// TIA Portal project "MCP_RB001002" (V15.1) (continued)
   SendWChar[1891] := WCHAR#' ';
   SendWChar[1892] := WCHAR#' ';
   SendWChar[1893] := WCHAR#' ';
   SendWChar[1894] := WCHAR#' ';
   SendWChar[1895] := WCHAR#' ';
   SendWChar[1896] := WCHAR#' ';
   SendWChar[1897] := WCHAR#' ';
   SendWChar[1898] := WCHAR#' ';
   SendWChar[1899] := WCHAR#' ';
   SendWChar[1900] := WCHAR#' ';
   SendWChar[1901] := WCHAR#' ';
   SendWChar[1902] := WCHAR#' ';
   SendWChar[1903] := WCHAR#' ';
   SendWChar[1904] := WCHAR#' ';
   SendWChar[1905] := WCHAR#' ';
   SendWChar[1906] := WCHAR#' ';
   SendWChar[1907] := WCHAR#' ';
   SendWChar[1908] := WCHAR#' ';
   SendWChar[1909] := WCHAR#' ';
   SendWChar[1910] := WCHAR#' ';
   SendWChar[1911] := WCHAR#' ';
   SendWChar[1912] := WCHAR#' ';
   SendWChar[1913] := WCHAR#' ';
   SendWChar[1914] := WCHAR#' ';
   SendWChar[1915] := WCHAR#' ';
   SendWChar[1916] := WCHAR#' ';
   SendWChar[1917] := WCHAR#' ';
   SendWChar[1918] := WCHAR#' ';
   SendWChar[1919] := WCHAR#' ';
   SendWChar[1920] := WCHAR#' ';
   SendWChar[1921] := WCHAR#' ';
   SendWChar[1922] := WCHAR#' ';
   SendWChar[1923] := WCHAR#' ';
   SendWChar[1924] := WCHAR#' ';
   SendWChar[1925] := WCHAR#' ';
   SendWChar[1926] := WCHAR#' ';
   SendWChar[1927] := WCHAR#' ';
   SendWChar[1928] := WCHAR#' ';
   SendWChar[1929] := WCHAR#' ';
   SendWChar[1930] := WCHAR#' ';
   SendWChar[1931] := WCHAR#' ';
   SendWChar[1932] := WCHAR#' ';
   SendWChar[1933] := WCHAR#' ';
   SendWChar[1934] := WCHAR#' ';
   SendWChar[1935] := WCHAR#' ';
   SendWChar[1936] := WCHAR#' ';
   SendWChar[1937] := WCHAR#' ';
   SendWChar[1938] := WCHAR#' ';
   SendWChar[1939] := WCHAR#' ';
   SendWChar[1940] := WCHAR#' ';
   SendWChar[1941] := WCHAR#' ';
   SendWChar[1942] := WCHAR#' ';
   SendWChar[1943] := WCHAR#' ';
   SendWChar[1944] := WCHAR#' ';
   SendWChar[1945] := WCHAR#' ';
   SendWChar[1946] := WCHAR#' ';
   SendWChar[1947] := WCHAR#' ';
   SendWChar[1948] := WCHAR#' ';
   SendWChar[1949] := WCHAR#' ';
   SendWChar[1950] := WCHAR#' ';
   SendWChar[1951] := WCHAR#' ';
   SendWChar[1952] := WCHAR#' ';
   SendWChar[1953] := WCHAR#' ';
   SendWChar[1954] := WCHAR#' ';
   SendWChar[1955] := WCHAR#' ';
   SendWChar[1956] := WCHAR#' ';
   SendWChar[1957] := WCHAR#' ';
   SendWChar[1958] := WCHAR#' ';
   SendWChar[1959] := WCHAR#' ';
   SendWChar[1960] := WCHAR#' ';
   SendWChar[1961] := WCHAR#' ';
   SendWChar[1962] := WCHAR#' ';
   SendWChar[1963] := WCHAR#' ';
   SendWChar[1964] := WCHAR#' ';
   SendWChar[1965] := WCHAR#' ';
   SendWChar[1966] := WCHAR#' ';
   SendWChar[1967] := WCHAR#' ';
   SendWChar[1968] := WCHAR#' ';
   SendWChar[1969] := WCHAR#' ';
   SendWChar[1970] := WCHAR#' ';
   SendWChar[1971] := WCHAR#' ';
   SendWChar[1972] := WCHAR#' ';
   SendWChar[1973] := WCHAR#' ';
   SendWChar[1974] := WCHAR#' ';
   SendWChar[1975] := WCHAR#' ';
   SendWChar[1976] := WCHAR#' ';
   SendWChar[1977] := WCHAR#' ';
   SendWChar[1978] := WCHAR#' ';
   SendWChar[1979] := WCHAR#' ';
   SendWChar[1980] := WCHAR#' ';
   SendWChar[1981] := WCHAR#' ';
   SendWChar[1982] := WCHAR#' ';
   SendWChar[1983] := WCHAR#' ';
   SendWChar[1984] := WCHAR#' ';
   SendWChar[1985] := WCHAR#' ';
   SendWChar[1986] := WCHAR#' ';
   SendWChar[1987] := WCHAR#' ';
   SendWChar[1988] := WCHAR#' ';
   SendWChar[1989] := WCHAR#' ';
   SendWChar[1990] := WCHAR#' ';
   SendWChar[1991] := WCHAR#' ';
   SendWChar[1992] := WCHAR#' ';
   SendWChar[1993] := WCHAR#' ';
   SendWChar[1994] := WCHAR#' ';
   SendWChar[1995] := WCHAR#' ';
   SendWChar[1996] := WCHAR#' ';
   SendWChar[1997] := WCHAR#' ';
   SendWChar[1998] := WCHAR#' ';
   SendWChar[1999] := WCHAR#' ';
   SendWChar[2000] := WCHAR#' ';
   SendWChar[2001] := WCHAR#' ';
   SendWChar[2002] := WCHAR#' ';
   SendWChar[2003] := WCHAR#' ';
   SendWChar[2004] := WCHAR#' ';
   SendWChar[2005] := WCHAR#' ';
   SendWChar[2006] := WCHAR#' ';
   SendWChar[2007] := WCHAR#' ';
   SendWChar[2008] := WCHAR#' ';
   SendWChar[2009] := WCHAR#' ';
   SendWChar[2010] := WCHAR#' ';
   SendWChar[2011] := WCHAR#' ';
   SendWChar[2012] := WCHAR#' ';
   SendWChar[2013] := WCHAR#' ';
   SendWChar[2014] := WCHAR#' ';
   SendWChar[2015] := WCHAR#' ';
   SendWChar[2016] := WCHAR#' ';
   SendWChar[2017] := WCHAR#' ';
   SendWChar[2018] := WCHAR#' ';
   SendWChar[2019] := WCHAR#' ';
   SendWChar[2020] := WCHAR#' ';
   SendWChar[2021] := WCHAR#' ';
   SendWChar[2022] := WCHAR#' ';
   SendWChar[2023] := WCHAR#' ';
   SendWChar[2024] := WCHAR#' ';
   SendWChar[2025] := WCHAR#' ';
   SendWChar[2026] := WCHAR#' ';
   SendWChar[2027] := WCHAR#' ';
   SendWChar[2028] := WCHAR#' ';
   SendWChar[2029] := WCHAR#' ';
   SendWChar[2030] := WCHAR#' ';
   SendWChar[2031] := WCHAR#' ';
   SendWChar[2032] := WCHAR#' ';
   SendWChar[2033] := WCHAR#' ';
   SendWChar[2034] := WCHAR#' ';
   SendWChar[2035] := WCHAR#' ';
   SendWChar[2036] := WCHAR#' ';
   SendWChar[2037] := WCHAR#' ';
   SendWChar[2038] := WCHAR#' ';
   SendWChar[2039] := WCHAR#' ';
   SendWChar[2040] := WCHAR#' ';
   SendWChar[2041] := WCHAR#' ';
   SendWChar[2042] := WCHAR#' ';
   SendWChar[2043] := WCHAR#' ';
   SendWChar[2044] := WCHAR#' ';
   SendWChar[2045] := WCHAR#' ';
   SendWChar[2046] := WCHAR#' ';
   SendWChar[2047] := WCHAR#' ';
   SendWChar[2048] := WCHAR#' ';
END_DATA_BLOCK

DATA_BLOCK "uMySQL_Use_DB"   // DB902
{ S7_Optimized_Access := 'TRUE' }
VERSION : 0.1
// stored: InstanceOfName uMySQL_Use
"uMySQL_Use"
BEGIN
END_DATA_BLOCK

DATA_BLOCK "uMySQL_Command_DB"   // DB903
{ S7_Optimized_Access := 'TRUE' }
VERSION : 0.1
// stored: InstanceOfName uMySQL_Command
"uMySQL_Command"
BEGIN
END_DATA_BLOCK

DATA_BLOCK "uMySQL_Query_DB"   // DB904
{ S7_Optimized_Access := 'TRUE' }
VERSION : 0.1
// stored: InstanceOfName uMySQL_Query
"uMySQL_Query"
BEGIN
END_DATA_BLOCK

// folder: (top level)

FUNCTION_BLOCK "温控相机解码"   // FB410, LAD
{ S7_Optimized_Access := 'TRUE' }
VERSION : 0.1
   VAR RETAIN
      Connparm : TCON_IP_v4;
   END_VAR
   VAR
      TRCV_C_Instance : TRCV_C;
      RECV_Data : Array[0..1023] of Byte;
   END_VAR
   // Connparm.InterfaceId := 64;
   // Connparm.ID := 16#65;
   // Connparm.ActiveEstablished := false;
   // Connparm.LocalPort := 9840;
BEGIN

REGION Network 1
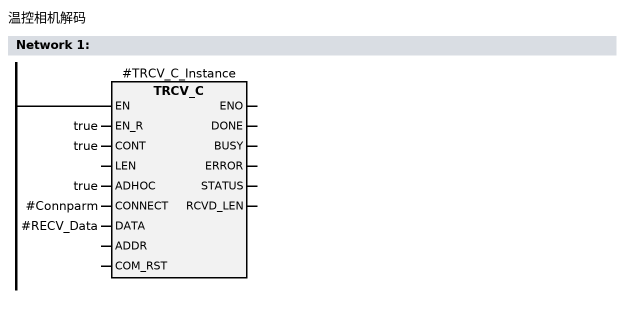
   #TRCV_C_Instance(EN_R := true, CONT := true, ADHOC := true, CONNECT := #Connparm, DATA := #RECV_Data);   // TRCV_C
END_REGION
END_FUNCTION_BLOCK

FUNCTION "精炼机数据处理" : Void   // FC100, LAD
{ S7_Optimized_Access := 'TRUE' }
VERSION : 0.1
   VAR_TEMP   // added for the SCL form of the ladder/FBD networks
      _w1 : Bool;
   END_VAR
BEGIN

REGION Network 1
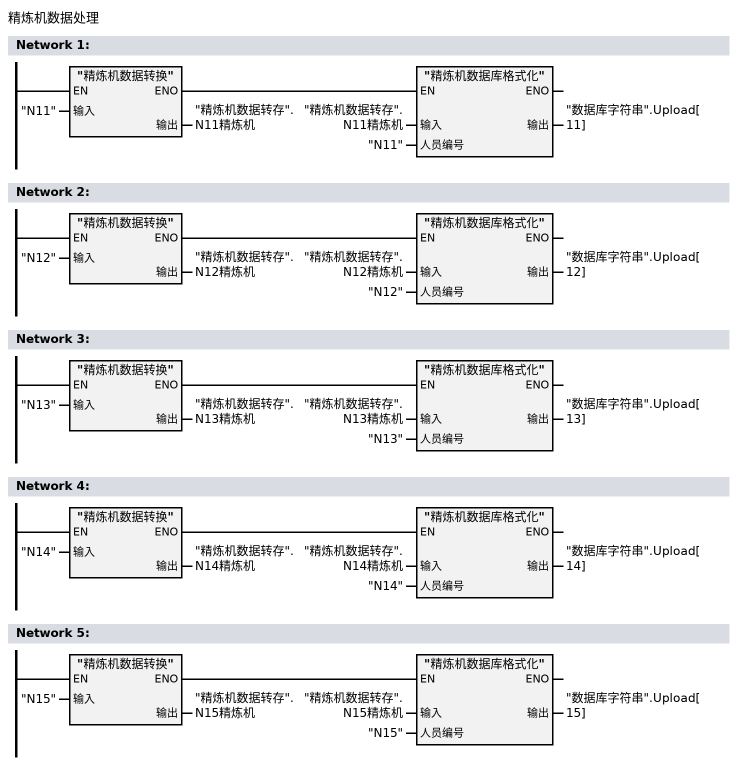
   RUNG wire#powerrail
      "精炼机数据转换"(输入 := "N11", 输出 => "精炼机数据转存".N11精炼机)
      "精炼机数据库格式化"(输入 := "精炼机数据转存".N11精炼机, 人员编号 := "N11", 输出 => "数据库字符串".Upload[11])
   END_RUNG
   // the same network as SCL:
   "精炼机数据转换"(输入 := "N11", 输出 => "精炼机数据转存".N11精炼机, ENO => #_w1);
   IF #_w1 THEN "精炼机数据库格式化"(输入 := "精炼机数据转存".N11精炼机, 人员编号 := "N11", 输出 => "数据库字符串".Upload[11]); END_IF;
END_REGION

REGION Network 2
   RUNG wire#powerrail
      "精炼机数据转换"(输入 := "N12", 输出 => "精炼机数据转存".N12精炼机)
      "精炼机数据库格式化"(输入 := "精炼机数据转存".N12精炼机, 人员编号 := "N12", 输出 => "数据库字符串".Upload[12])
   END_RUNG
   // the same network as SCL:
   "精炼机数据转换"(输入 := "N12", 输出 => "精炼机数据转存".N12精炼机, ENO => #_w1);
   IF #_w1 THEN "精炼机数据库格式化"(输入 := "精炼机数据转存".N12精炼机, 人员编号 := "N12", 输出 => "数据库字符串".Upload[12]); END_IF;
END_REGION

REGION Network 3
   RUNG wire#powerrail
      "精炼机数据转换"(输入 := "N13", 输出 => "精炼机数据转存".N13精炼机)
      "精炼机数据库格式化"(输入 := "精炼机数据转存".N13精炼机, 人员编号 := "N13", 输出 => "数据库字符串".Upload[13])
   END_RUNG
   // the same network as SCL:
   "精炼机数据转换"(输入 := "N13", 输出 => "精炼机数据转存".N13精炼机, ENO => #_w1);
   IF #_w1 THEN "精炼机数据库格式化"(输入 := "精炼机数据转存".N13精炼机, 人员编号 := "N13", 输出 => "数据库字符串".Upload[13]); END_IF;
END_REGION

REGION Network 4
   RUNG wire#powerrail
      "精炼机数据转换"(输入 := "N14", 输出 => "精炼机数据转存".N14精炼机)
      "精炼机数据库格式化"(输入 := "精炼机数据转存".N14精炼机, 人员编号 := "N14", 输出 => "数据库字符串".Upload[14])
   END_RUNG
   // the same network as SCL:
   "精炼机数据转换"(输入 := "N14", 输出 => "精炼机数据转存".N14精炼机, ENO => #_w1);
   IF #_w1 THEN "精炼机数据库格式化"(输入 := "精炼机数据转存".N14精炼机, 人员编号 := "N14", 输出 => "数据库字符串".Upload[14]); END_IF;
END_REGION

REGION Network 5
   RUNG wire#powerrail
      "精炼机数据转换"(输入 := "N15", 输出 => "精炼机数据转存".N15精炼机)
      "精炼机数据库格式化"(输入 := "精炼机数据转存".N15精炼机, 人员编号 := "N15", 输出 => "数据库字符串".Upload[15])
   END_RUNG
   // the same network as SCL:
   "精炼机数据转换"(输入 := "N15", 输出 => "精炼机数据转存".N15精炼机, ENO => #_w1);
   IF #_w1 THEN "精炼机数据库格式化"(输入 := "精炼机数据转存".N15精炼机, 人员编号 := "N15", 输出 => "数据库字符串".Upload[15]); END_IF;
END_REGION
END_FUNCTION

FUNCTION "SWP_Word" : WChar   // FC108, SCL
{ S7_Optimized_Access := 'TRUE' }
VERSION : 0.1
   VAR_INPUT
      IW : Word;
   END_VAR
   VAR_TEMP
      TempWord : Word;
   END_VAR
BEGIN
   #TempWord.%B0 := #IW.%B1;
   #TempWord.%B1 := #IW.%B0;
   #SWP_Word := WORD_TO_WCHAR(#TempWord);
END_FUNCTION

FUNCTION "SWP_Lreal" : Real   // FC109, SCL
{ S7_Optimized_Access := 'TRUE' }
VERSION : 0.1
   VAR_INPUT
      ID : Real;
   END_VAR
   VAR_TEMP
      TempWord : DWord;
      TempDword : DWord;
   END_VAR
BEGIN
   #TempDword := REAL_TO_DWORD(#ID);
   #TempWord.%B0 := #TempDword.%B2;
   #TempWord.%B1 := #TempDword.%B3;
   #TempWord.%B2 := #TempDword.%B0;
   #TempWord.%B3 := #TempDword.%B1;
   #SWP_Lreal := DWORD_TO_REAL(#TempWord);
END_FUNCTION

FUNCTION "精炼机数据转换" : Void   // FC110, SCL
{ S7_Optimized_Access := 'TRUE' }
VERSION : 0.1
   VAR_INPUT
      输入 : "精炼机";
   END_VAR
   VAR_OUTPUT
      输出 : "精炼机上传";
   END_VAR
BEGIN
   #输出.左前辊温度 := "SWP_Lreal"(#输入.左前辊温度);
   #输出.右前辊温度 := "SWP_Lreal"(#输入.右前辊温度);
   #输出.左后辊温度 :="SWP_Lreal"( #输入.左后辊温度);
   #输出.右后辊温度 :="SWP_Lreal"( #输入.右后辊温度);
   #输出.左间隙 :="SWP_Lreal"( #输入.左间隙) ;
   #输出.右间隙 :="SWP_Lreal"( #输入.右间隙);
   #输出.滚筒电机电流 := "SWP_Lreal"(#输入.滚筒电机电流);
   #输出.滚筒电机频率 :="SWP_Lreal"( #输入.滚筒电机频率);
   #输出.滚筒电机功率 :="SWP_Lreal"( #输入.滚筒电机功率);
   #输出.滚筒电机电度 :="SWP_DINT"( #输入.滚筒电机电度);
   #输出.滚筒电机计时 :="SWP_DINT"( #输入.滚筒电机计时) ;
   #输出.环境温度 := "通用数据采集".环境温度;//"SWP_Lreal"( #输入.环境温度);
   #输出.环境湿度 := "通用数据采集".环境湿度;//"SWP_Lreal"( #输入.环境湿度);
   #输出.胶温 :="SWP_Lreal"( #输入.胶温);
   #输出.开关量汇总 :="SWP_DINT"( #输入.开关量汇总);

   #输出.当前任务编号[0] := "SWP_Word"(#输入.当前任务编号[0]);
   #输出.当前任务编号[1] := "SWP_Word"(#输入.当前任务编号[1]);
   #输出.当前任务编号[2] := "SWP_Word"(#输入.当前任务编号[2]);
   #输出.当前任务编号[3] := "SWP_Word"(#输入.当前任务编号[3]);
   #输出.当前任务编号[4] := "SWP_Word"(#输入.当前任务编号[4]);
   #输出.当前任务编号[5] := "SWP_Word"(#输入.当前任务编号[5]);
   #输出.当前任务编号[6] := "SWP_Word"(#输入.当前任务编号[6]);
   #输出.当前任务编号[7] := "SWP_Word"(#输入.当前任务编号[7]);
   #输出.当前任务编号[8] := "SWP_Word"(#输入.当前任务编号[8]);
   #输出.当前任务编号[9] := "SWP_Word"(#输入.当前任务编号[9]);
   #输出.当前人员编号[0] := "SWP_Word"(#输入.当前人员编号[0]);
   #输出.当前人员编号[1] := "SWP_Word"(#输入.当前人员编号[1]);
   #输出.当前人员编号[2] := "SWP_Word"(#输入.当前人员编号[2]);
   #输出.当前人员编号[3] := "SWP_Word"(#输入.当前人员编号[3]);
   #输出.当前人员编号[4] := "SWP_Word"(#输入.当前人员编号[4]);
   #输出.当前人员编号[5] := "SWP_Word"(#输入.当前人员编号[5]);
   #输出.当前人员编号[6] := "SWP_Word"(#输入.当前人员编号[6]);
   #输出.当前人员编号[7] := "SWP_Word"(#输入.当前人员编号[7]);
   #输出.当前人员编号[8] := "SWP_Word"(#输入.当前人员编号[8]);
   #输出.当前人员编号[9] := "SWP_Word"(#输入.当前任务编号[9]);
END_FUNCTION

FUNCTION "SWP_DINT" : DInt   // FC111, SCL
{ S7_Optimized_Access := 'TRUE' }
VERSION : 0.1
   VAR_INPUT
      ID : DInt;
   END_VAR
   VAR_TEMP
      TempWord : DWord;
      TempDword : DWord;
   END_VAR
BEGIN
   #TempDword := DINT_TO_DWORD(#ID);
   #TempWord.%B0 := #TempDword.%B2;
   #TempWord.%B1 := #TempDword.%B3;
   #TempWord.%B2 := #TempDword.%B0;
   #TempWord.%B3 := #TempDword.%B1;
   #SWP_DINT := DWORD_TO_DINT(#TempWord);
END_FUNCTION

FUNCTION "两点校正输入" : Void   // FC168, SCL
{ S7_Optimized_Access := 'TRUE' }
VERSION : 0.1
   VAR_INPUT
      Max : Real;
      PIW : Word;
      Min : Real;
      Full : Int;
      Zero : Int;
   END_VAR
   VAR_OUTPUT
      RealValue : Real;
      Error : Bool;
   END_VAR
BEGIN
   #RealValue := ((#Max - #Min) / INT_TO_REAL(#Full - #Zero)) * INT_TO_REAL(WORD_TO_INT(#PIW) - #Zero) + #Min;
   #RealValue := LIMIT(MN := #Min, IN := #RealValue, MX := #Max);
   IF #PIW = 16#7fff OR #PIW = 16#8000 THEN
       #Error := true;
   END_IF;
END_FUNCTION

FUNCTION "通用数据处理" : Void   // FC200, LAD
{ S7_Optimized_Access := 'TRUE' }
VERSION : 0.1
   VAR_TEMP   // added for the SCL form of the ladder/FBD networks
      _w1 : Bool;
      _w2 : Bool;
   END_VAR
BEGIN

REGION Network 1
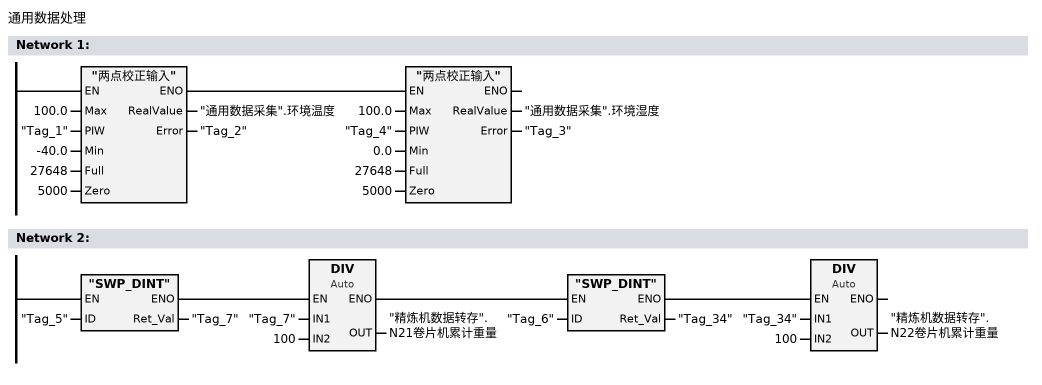
   RUNG wire#powerrail
      "两点校正输入"(Max := 100.0, PIW := "Tag_1", Min := -40.0, Full := 27648, Zero := 5000, RealValue => "通用数据采集".环境温度, Error => "Tag_2")
      "两点校正输入"(Max := 100.0, PIW := "Tag_4", Min := 0.0, Full := 27648, Zero := 5000, RealValue => "通用数据采集".环境湿度, Error => "Tag_3")
   END_RUNG
   // the same network as SCL:
   "两点校正输入"(Max := 100.0,
            PIW := "Tag_1",
            Min := -40.0,
            Full := 27648,
            Zero := 5000,
            RealValue => "通用数据采集".环境温度,
            Error => "Tag_2",
            ENO => #_w1);
   IF #_w1 THEN
       "两点校正输入"(Max := 100.0,
                PIW := "Tag_4",
                Min := 0.0,
                Full := 27648,
                Zero := 5000,
                RealValue => "通用数据采集".环境湿度,
                Error => "Tag_3");
   END_IF;
END_REGION

REGION Network 2
   RUNG wire#powerrail
      "SWP_DINT"(ID := "Tag_5", Ret_Val => "Tag_7")
      Div(in1 := "Tag_7", in2 := 100, out => "精炼机数据转存".N21卷片机累计重量)
      "SWP_DINT"(ID := "Tag_6", Ret_Val => "Tag_34")
      Div(in1 := "Tag_34", in2 := 100, out => "精炼机数据转存".N22卷片机累计重量)
   END_RUNG
   // the same network as SCL:
   "Tag_7" := "SWP_DINT"(ID := "Tag_5", ENO => #_w1);
   IF #_w1 THEN "精炼机数据转存".N21卷片机累计重量 := "Tag_7" / 100; END_IF;
   "Tag_34" := "SWP_DINT"(EN := #_w1, ID := "Tag_6", ENO => #_w2);
   IF #_w2 THEN "精炼机数据转存".N22卷片机累计重量 := "Tag_34" / 100; END_IF;
END_REGION
END_FUNCTION

FUNCTION "温控相机通信" : Void   // FC400, LAD
{ S7_Optimized_Access := 'TRUE' }
VERSION : 0.1
BEGIN

REGION Network 1
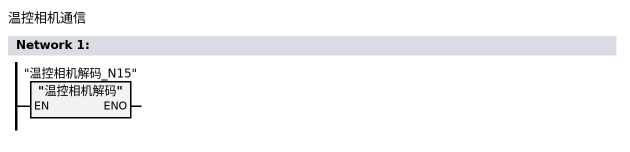
   RUNG wire#powerrail
      "温控相机解码_N15"()
   END_RUNG
   // the same network as SCL:
   "温控相机解码_N15"();   // "温控相机解码"
END_REGION
END_FUNCTION

ORGANIZATION_BLOCK "Main"   // OB1, LAD, ProgramCycle
TITLE = "Main Program Sweep (Cycle)"
{ S7_Optimized_Access := 'TRUE' }
VERSION : 0.1
   VAR_INPUT
      Initial_Call : Bool;   // Initial call of this OB
      Remanence : Bool;   // =True, if remanent data are available
   END_VAR
BEGIN

REGION Network 1
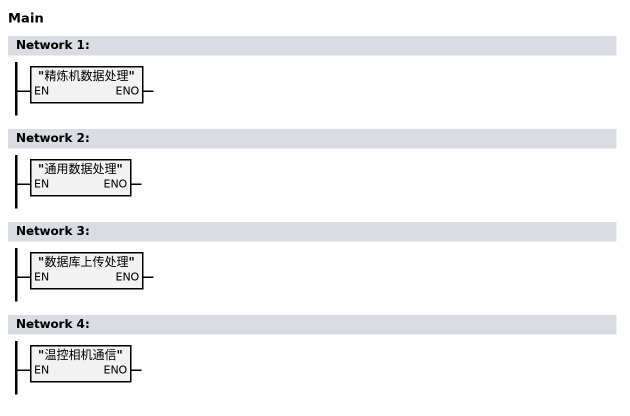
   RUNG wire#powerrail
      "精炼机数据处理"()
   END_RUNG
   // the same network as SCL:
   "精炼机数据处理"();
END_REGION

REGION Network 2
   RUNG wire#powerrail
      "通用数据处理"()
   END_RUNG
   // the same network as SCL:
   "通用数据处理"();
END_REGION

REGION Network 3
   RUNG wire#powerrail
      "数据库上传处理"()
   END_RUNG
   // the same network as SCL:
   "数据库上传处理"();
END_REGION

REGION Network 4
   RUNG wire#powerrail
      "温控相机通信"()
   END_RUNG
   // the same network as SCL:
   "温控相机通信"();
END_REGION
END_ORGANIZATION_BLOCK

// folder: 存数据库

FUNCTION "数据库上传处理" : Void   // FC300, LAD
{ S7_Optimized_Access := 'TRUE' }
VERSION : 0.1
BEGIN

REGION Network 1
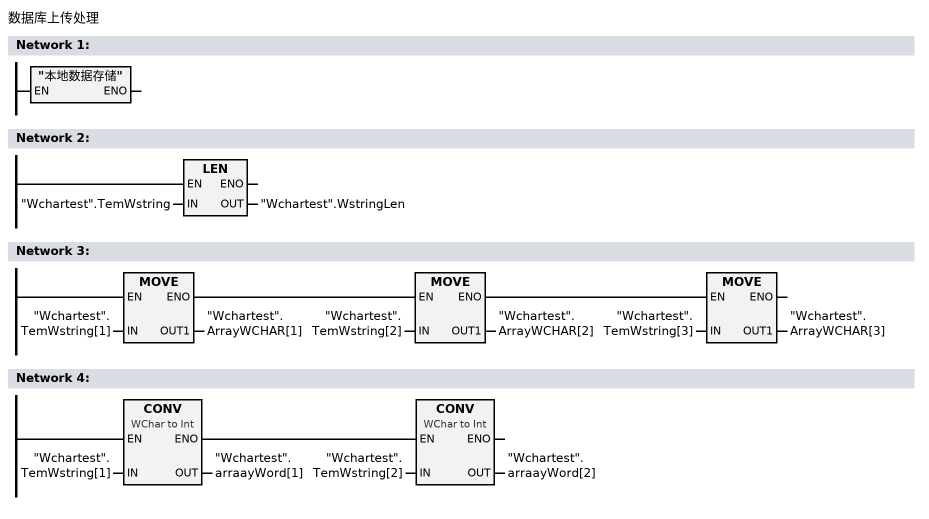
   RUNG wire#powerrail
      "本地数据存储"()
   END_RUNG
   // the same network as SCL:
   "本地数据存储"();
END_REGION

REGION Network 2
   "Wchartest".WstringLen := LEN(IN := "Wchartest".TemWstring);
END_REGION

REGION Network 3
   RUNG wire#powerrail
      Move(in := "Wchartest".TemWstring[1], out1 => "Wchartest".ArrayWCHAR[1])
      Move(in := "Wchartest".TemWstring[2], out1 => "Wchartest".ArrayWCHAR[2])
      Move(in := "Wchartest".TemWstring[3], out1 => "Wchartest".ArrayWCHAR[3])
   END_RUNG
   // the same network as SCL:
   "Wchartest".ArrayWCHAR[1] := "Wchartest".TemWstring[1];
   "Wchartest".ArrayWCHAR[2] := "Wchartest".TemWstring[2];
   "Wchartest".ArrayWCHAR[3] := "Wchartest".TemWstring[3];
END_REGION

REGION Network 4
   RUNG wire#powerrail
      { S7_Templates := "[SrcType := WChar, DestType := Int]" } Convert(in := "Wchartest".TemWstring[1], out => "Wchartest".arraayWord[1])
      { S7_Templates := "[SrcType := WChar, DestType := Int]" } Convert(in := "Wchartest".TemWstring[2], out => "Wchartest".arraayWord[2])
   END_RUNG
   // the same network as SCL:
   "Wchartest".arraayWord[1] := WCHAR_TO_INT("Wchartest".TemWstring[1]);
   "Wchartest".arraayWord[2] := WCHAR_TO_INT("Wchartest".TemWstring[2]);
END_REGION
END_FUNCTION

FUNCTION "精炼机数据库格式化" : Void   // FC311, SCL
{ S7_Optimized_Access := 'TRUE' }
VERSION : 0.1
   VAR_INPUT
      输入 : "精炼机上传";
      人员编号 : "精炼机";
   END_VAR
   VAR_OUTPUT
      输出 : "精炼机数据库";
   END_VAR
BEGIN
   #输出.左前辊温度 := #输入.左前辊温度;
   #输出.右前辊温度 := #输入.右前辊温度;
   #输出.左后辊温度 := #输入.左后辊温度;
   #输出.右后辊温度 := #输入.右后辊温度;
   #输出.左间隙 := #输入.左间隙;
   #输出.右间隙 := #输入.右间隙;
   #输出.滚筒电机电流 := #输入.滚筒电机电流;
   #输出.滚筒电机频率 := #输入.滚筒电机频率;
   #输出.滚筒电机功率 := #输入.滚筒电机功率;
   #输出.滚筒电机电度 := #输入.滚筒电机电度;
   #输出.滚筒电机计时 := #输入.滚筒电机计时;
   #输出.环境温度 := #输入.环境温度;
   #输出.环境湿度 := #输入.环境湿度;
   #输出.胶温 := #输入.胶温;
   #输出.开关量汇总 := #输入.开关量汇总;
   Chars_TO_Strg(Chars:=#人员编号.当前任务编号,
                             pChars:=0,
                             Cnt:=16,
                             Strg=>#输出.当前任务编号);
               Chars_TO_Strg(Chars := #人员编号.当前人员编号,
                             pChars := 0,
                             Cnt := 16,
                             Strg => #输出.当前人员编号);
END_FUNCTION

FUNCTION "轮训写入数据" : Void   // FC321, LAD
{ S7_Optimized_Access := 'TRUE' }
VERSION : 0.1
BEGIN

REGION Network 1
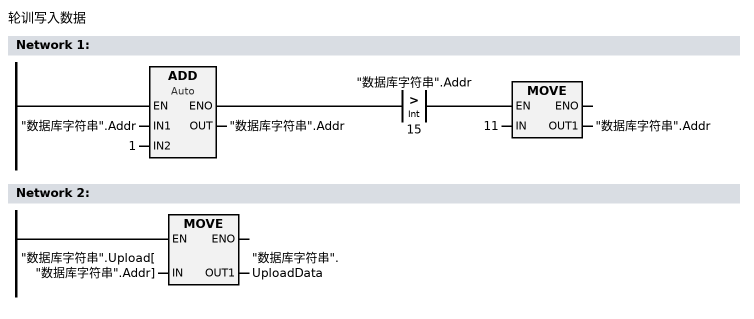
   RUNG wire#powerrail
      Add(in1 := "数据库字符串".Addr, in2 := 1, out => "数据库字符串".Addr)
      { S7_Templates := "SrcType := Int" } GT_Contact(in1 := "数据库字符串".Addr, in2 := 15)
      Move(in := 11, out1 => "数据库字符串".Addr)
   END_RUNG
   // the same network as SCL:
   "数据库字符串".Addr := "数据库字符串".Addr + 1;
   IF "数据库字符串".Addr > 15 THEN "数据库字符串".Addr := 11; END_IF;
END_REGION

REGION Network 2
   RUNG wire#powerrail
      Move(in := "数据库字符串".Upload["数据库字符串".Addr], out1 => "数据库字符串".UploadData)
   END_RUNG
   // the same network as SCL:
   "数据库字符串".UploadData := "数据库字符串".Upload["数据库字符串".Addr];
END_REGION
END_FUNCTION

FUNCTION "本地数据存储" : Void   // FC900, LAD
{ S7_Optimized_Access := 'TRUE' }
VERSION : 0.1
   VAR_TEMP   // added for the SCL form of the ladder/FBD networks
      _w1 : Bool;
      _w2 : Bool;
   END_VAR
BEGIN

REGION Network 1: 连接数据库
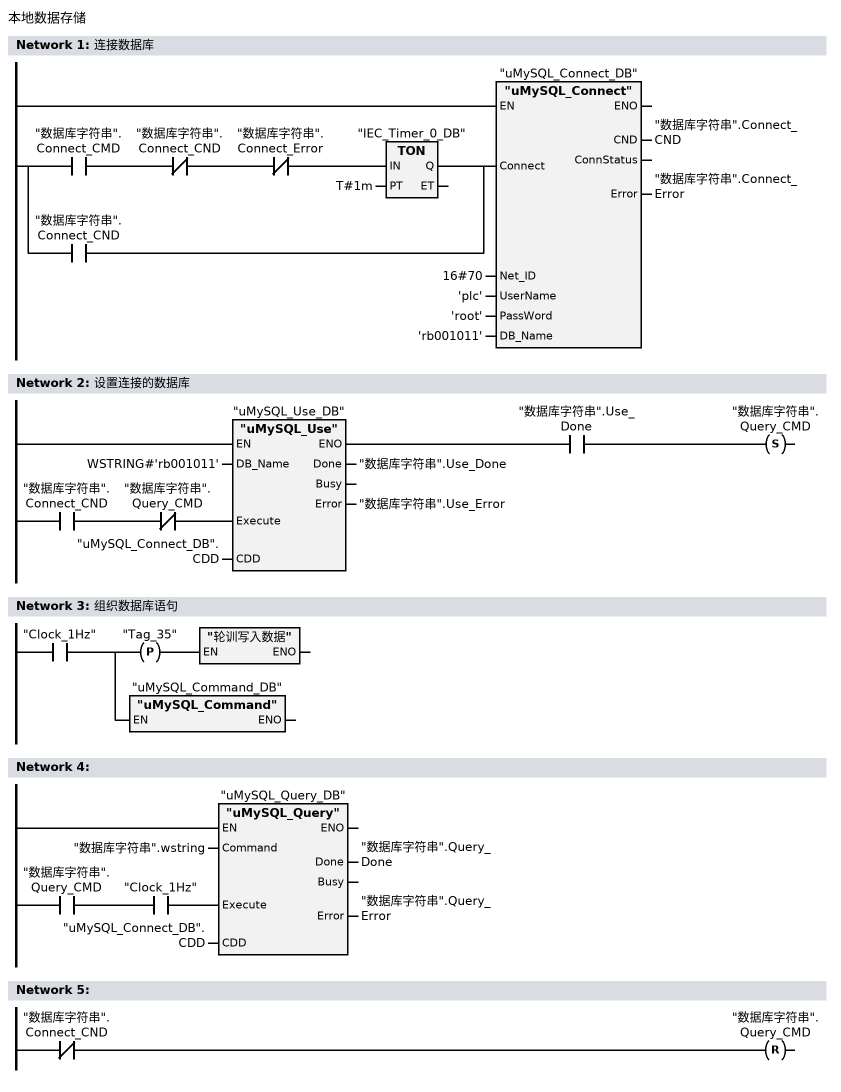
   "IEC_Timer_0_DB".TON(IN := "数据库字符串".Connect_CMD AND NOT "数据库字符串".Connect_CND AND NOT "数据库字符串".Connect_Error,
                        PT := T#1m);
   "uMySQL_Connect_DB"(Connect := "IEC_Timer_0_DB".Q OR "数据库字符串".Connect_CND,   // "uMySQL_Connect"
                       Net_ID := 16#70,
                       UserName := 'plc',
                       PassWord := 'root',
                       DB_Name := 'rb001011',
                       CND => "数据库字符串".Connect_CND,
                       Error => "数据库字符串".Connect_Error);
END_REGION

REGION Network 2: 设置连接的数据库
   RUNG wire#powerrail
      "uMySQL_Use_DB"(Execute := wire#w1, DB_Name := WSTRING#'rb001011', CDD := "uMySQL_Connect_DB".CDD, Done => "数据库字符串".Use_Done, Busy =>, Error => "数据库字符串".Use_Error)
      Contact( "数据库字符串".Use_Done )
      S_Coil( "数据库字符串".Query_CMD )
   END_RUNG
   RUNG wire#powerrail
      Contact( "数据库字符串".Connect_CND )
      I_Contact( "数据库字符串".Query_CMD )
   END_RUNG wire#w1
   // the same network as SCL:
   "uMySQL_Use_DB"(DB_Name := WSTRING#'rb001011',   // "uMySQL_Use"
                   Execute := "数据库字符串".Connect_CND AND NOT "数据库字符串".Query_CMD,
                   CDD := "uMySQL_Connect_DB".CDD,
                   Done => "数据库字符串".Use_Done,
                   Error => "数据库字符串".Use_Error,
                   ENO => #_w1);
   IF #_w1 AND "数据库字符串".Use_Done THEN "数据库字符串".Query_CMD := TRUE; END_IF;
END_REGION

REGION Network 3: 组织数据库语句
   RUNG wire#powerrail
      Contact( "Clock_1Hz" )
      wire#w1
      P_Trig( "Tag_35" )
      "轮训写入数据"()
   END_RUNG
   RUNG wire#w1
      "uMySQL_Command_DB"()
   END_RUNG
   // the same network as SCL:
   #_w1 := "Clock_1Hz" AND NOT "Tag_35";   // rising edge
   "Tag_35" := "Clock_1Hz";
   #_w2 := "Clock_1Hz";
   IF #_w1 THEN "轮训写入数据"(); END_IF;
   IF #_w2 THEN
       "uMySQL_Command_DB"();   // "uMySQL_Command"
   END_IF;
END_REGION

REGION Network 4
   RUNG wire#powerrail
      "uMySQL_Query_DB"(Execute := wire#w1, Command := "数据库字符串".wstring, CDD := "uMySQL_Connect_DB".CDD, Done => "数据库字符串".Query_Done, Busy =>, Error => "数据库字符串".Query_Error)
   END_RUNG
   RUNG wire#powerrail
      Contact( "数据库字符串".Query_CMD )
      Contact( "Clock_1Hz" )
   END_RUNG wire#w1
   // the same network as SCL:
   "uMySQL_Query_DB"(Command := "数据库字符串".wstring,   // "uMySQL_Query"
                     Execute := "数据库字符串".Query_CMD AND "Clock_1Hz",
                     CDD := "uMySQL_Connect_DB".CDD,
                     Done => "数据库字符串".Query_Done,
                     Error => "数据库字符串".Query_Error);
END_REGION

REGION Network 5
   RUNG wire#powerrail
      I_Contact( "数据库字符串".Connect_CND )
      R_Coil( "数据库字符串".Query_CMD )
   END_RUNG
   // the same network as SCL:
   IF NOT "数据库字符串".Connect_CND THEN "数据库字符串".Query_CMD := FALSE; END_IF;
END_REGION

REGION Network 6: 每次PLC上电，流水号自加
END_REGION
END_FUNCTION

// folder: 存数据库/uMySQL

FUNCTION_BLOCK "uMySQL_Connect"   // FB3, SCL
{ S7_Optimized_Access := 'TRUE' }
VERSION : 0.1
   VAR_INPUT
      Connect : Bool;   // True:发起连接；False:断开连接 / 发起连接
      Net_ID : Conn_Ouc;   // 连接ID
      UserName : String := 'root';   // 数据库用户名
      PassWord : String := 'root';   // 数据库密码
      DB_Name : String := 'hist';   // 数据库名 / 数据库名称
   END_VAR
   VAR_OUTPUT
      CND : Bool;   // 连接成功
      ConnStatus : Byte;   // 连接状态
      Error : Bool;   // 错误
   END_VAR
   VAR
      IP : TCON_IP_v4;
      CDD : "uMySQL_CDD";   // 共用的数据库连接参数
      TempBool : Array[0..19] of Bool;
      REV_Buffer : Array[0..#MessageMaxLen] of Byte;
      SND_Buffer : Array[0..#MessageMaxLen] of Byte;
      NetConnect : TCON;
      NetRcv : TRCV;
      NetRcv_EN : Bool;
      NetRcv_Len : Int;
      NetRcv_Done : Bool;
      "Step" : Int;
      MessageLen : Int;   // 消息帧长度
      SaltLen : Int;   // 挑战随机数长度
      Server_Auth_PlugIn_Name : String;
      ServerVersion_StartNum : Int;
      ServerCapability_flag : DWord;
      SaltString : Array[0..49] of Byte;
      Client_CapabilityFlag : DWord := 16#8609;   // 客户端权能标志位
      Client_MaxLen : DWord;
      Calc_Encryption_SHA1 : "Calc_Encryption_SHA1";
      Temp_SHA1 : Array[0..19] of Byte;
      Temp_SHA_Arry : Array[0..55] of Byte;
      Temp_SHA_Arry_Num : UInt;
      Temp_SHA_Arry_Num_Int : Int;
      Temp_SHA1_2 : Array[0..19] of Byte;
      Temp_SHA1_3 : Array[0..19] of Byte;
      Token : Array[0..19] of Byte;
      NetDISCON : TDISCON;
      NetDiscon_EN : Bool;
      NetSend : TSEND;
      NetSend_EN : Bool;
      NetSend_Done : Bool;
      TDiag_Result : TDiag_Status;
      NetDiag : T_DIAG;
      NetDiag_EN : Bool;
      NetSendLen : Int;
      Timer_ON : TON_TIME;
      Timer_OFF : TON_TIME;
      Timer_Error : TON_TIME;
      NetSendEnd : TSEND;
      NetSendEnd_EN : Bool;
      NetSendEnd_Done : Bool;
      Command_Len : UInt;
      SendWChar : Array[0..2048] of WChar;
      Temp_CND : Bool;   // 连接成功
      Temp_ConnStatus : Byte;   // 连接状态
      Temp_NowNum : Int;
   END_VAR
   VAR_TEMP
      Temp_Dword : DWord;
      Temp_Index_i : Int;
      Temp_StrLen : Int;
   END_VAR
   VAR CONSTANT
      MessageMaxLen : DInt := 2048;   // 收发消息的最大长度
   END_VAR
   // IP.RemotePort := 3306;
   // IP.RemoteAddress.ADDR[4] := 16#A8;
   // IP.RemoteAddress.ADDR[3] := 16#1F;
   // IP.RemoteAddress.ADDR[2] := 16#A8;
   // IP.RemoteAddress.ADDR[1] := 16#C0;
   // IP.ActiveEstablished := true;
   // // CDD.Connect_OK : 数据库是否连接状态True:已连接；False :未连接
   // // CDD.Connect_ID : 连接ID，用于传递
   // // CDD.Connect_Sequence : 命令Sequence，用于传递
BEGIN


   (***********************************************************初始化数据******************************************************************)
   IF #Connect AND  #TempBool[0]=FALSE THEN
       #TempBool[0] := TRUE;
       #TempBool[1] := FALSE;
       #Step := 0;
       #CDD.Connect_ID := #Net_ID;
       #IP.ID := #Net_ID;
       #NetConnect.DONE := FALSE;
       #NetRcv_EN := TRUE;
       #NetDiscon_EN := FALSE;
       #NetSendEnd_EN := FALSE;
       ;
   END_IF;
   //#CDD.Recv_Done := FALSE;
   (***********************************************************断开连接******************************************************************)
   IF #Connect = FALSE AND #TempBool[1]=FALSE THEN
       #TempBool[0] := FALSE;
       #TempBool[1] := TRUE;
       //#NetRcv_EN := FALSE;
       #Step := 6;
   END_IF;


   #NetConnect(REQ:=#Connect,
               ID:=  #CDD.Connect_ID,
               CONNECT:=#IP);
   #NetRcv(EN_R:=#NetRcv_EN,
           ID:=#CDD.Connect_ID,
           LEN:=0,
           ADHOC:=TRUE,
           DATA:=#REV_Buffer);
   IF #NetRcv.NDR THEN
       #NetRcv_Done := TRUE;
       #NetRcv_Len := UDINT_TO_INT(#NetRcv.RCVD_LEN);
   END_IF;
   (***********************************************************处理流程******************************************************************)
   //#Step 0  发起连接
   //#Step 1 等待MySQL服务器发回来的数据
   //#Step 2 解码发回来的认证数据，并计算需要响应的数据放入Sendbuffer
   //#Step 3 开始发送并等待发送完成
   //#Step 4 发送完成等待返回认证结果
   //#Step 5 解析返回结果是否已经连接成功
   //#Step 6 申请断开连接

   CASE #Step OF
       0:  // 如果在等待服务器第一次连接
           IF #NetConnect.DONE THEN
               #Step := 1;
           END_IF;
       1:  // 连接并等待返回第一次握手数据
           IF     #NetRcv_Done  THEN
               #NetRcv_Done := FALSE;
               #Step := 2;
               #NetRcv_EN := FALSE;
               #NetRcv_Len := UDINT_TO_INT(#NetRcv.RCVD_LEN);
           END_IF;
       2:
           REGION MySQL_Auth_Packet
               #Temp_Dword.%B0 := #REV_Buffer[0];
               #Temp_Dword.%B1 := #REV_Buffer[1];
               #Temp_Dword.%B2 := #REV_Buffer[2];
               #Temp_Dword.%B3 := b#16#00;
               #MessageLen := DINT_TO_INT(DWORD_TO_DINT(#Temp_Dword)); //实际传输数据的字符长度
               #CDD.Connect_Sequence := BYTE_TO_INT(#REV_Buffer[3]); //传输的Sequence值

               #CDD.Server_Protocol_Version := BYTE_TO_INT(#REV_Buffer[4]); //MySQL服务器的协议版本号，当前大多为10(16#0A)
               #ServerVersion_StartNum := 5;
               WHILE #REV_Buffer[#ServerVersion_StartNum] <> b#16#00 DO//MySQL服务器的版本号，第5个字符开始，00结尾
                   #CDD.Server_Server_Version[#ServerVersion_StartNum-4] := #REV_Buffer[#ServerVersion_StartNum];
                   #ServerVersion_StartNum := #ServerVersion_StartNum + 1;
               END_WHILE;
               #ServerVersion_StartNum := #ServerVersion_StartNum + 1;//b#16#00是服务器版本号的结尾，要跳到下一个字节
               #ServerVersion_StartNum := #ServerVersion_StartNum + 4;//跳过服务器线程ID

               FOR #Temp_Index_i := 0 TO 7 DO
                   #SaltString[#Temp_Index_i] := #REV_Buffer[#ServerVersion_StartNum];//挑战字符串的前8个Byte
                   #ServerVersion_StartNum := #ServerVersion_StartNum + 1;
               END_FOR;
               #ServerVersion_StartNum := #ServerVersion_StartNum + 1;
               #ServerCapability_flag.%B3 := #REV_Buffer[#ServerVersion_StartNum];//权能标志位低-低字节
               #ServerVersion_StartNum := #ServerVersion_StartNum + 1;
               #ServerCapability_flag.%B2 := #REV_Buffer[#ServerVersion_StartNum];//权能标志位低-高字节
               #ServerVersion_StartNum := #ServerVersion_StartNum + 1;
               #CDD.Server_Character_Set := #REV_Buffer[#ServerVersion_StartNum]; //采用字符集
               #ServerVersion_StartNum := #ServerVersion_StartNum + 1;
               #ServerVersion_StartNum := #ServerVersion_StartNum + 2;
               #ServerCapability_flag.%B1 := #REV_Buffer[#ServerVersion_StartNum];//权能标志位高-低字节
               #ServerVersion_StartNum := #ServerVersion_StartNum + 1;
               #ServerCapability_flag.%B0 := #REV_Buffer[#ServerVersion_StartNum];//权能标志位高-高字节
               #ServerVersion_StartNum := #ServerVersion_StartNum + 1;
               #SaltLen := BYTE_TO_INT(#REV_Buffer[#ServerVersion_StartNum]) -1; //采用挑战随机数的数量
               #ServerVersion_StartNum := #ServerVersion_StartNum + 1;
               #ServerVersion_StartNum := #ServerVersion_StartNum + 10;//跳过保留的10个B#16#00
               FOR #Temp_Index_i := 0 TO #SaltLen - 9 DO   //去掉前面的8个数据，同时从0开始，所以-9
                   #SaltString[#Temp_Index_i + 8] := #REV_Buffer[#ServerVersion_StartNum];//挑战字符串的后面N个Byte
                   #ServerVersion_StartNum := #ServerVersion_StartNum + 1;
               END_FOR;
               #ServerVersion_StartNum := #ServerVersion_StartNum + 1;
               #Temp_Index_i := 0;
               WHILE #REV_Buffer[#ServerVersion_StartNum] <> b#16#00 DO//MySQL服务器的版本号，第5个字符开始，00结尾
                   #CDD.CLIENT_PLUGIN_AUTH[#Temp_Index_i+1] := #REV_Buffer[#ServerVersion_StartNum];
                   #ServerVersion_StartNum := #ServerVersion_StartNum + 1;
                   #Temp_Index_i := #Temp_Index_i + 1;
               END_WHILE;

